screen "41 BWT Ops" 1280x800, template "Template"
   TextField "Text field_60" at 920,365 size 100x30; Text 'GCU'
   GraphicIOField "Graphic I/O field_4" at 920,395 size 100x90; PictureList "GCU"
      ProcessValue <- "100_GCU_AUTO_SEQ_DB_RNG"
   TextField "Text field_70" at 930,485 size 80x25; Text 'Disabled'
   TextField "Text field_71" at 930,485 size 80x25; Text 'Enabled'
      Visibility <- "100_GCU_AUTO_SEQ_DB_RNG"
   Button "Button_4" at 910,355 size 120x170; TextOff 'Text'
      on Release: ActivateScreen("Inert Gas Conditioning Plant", 0)
   TextField "Text field_65" at 730,365 size 100x30; Text 'PGC'
   TextField "Text field_75" at 740,485 size 80x25; Text 'Disabled'
   TextField "Text field_76" at 740,485 size 80x25; Text 'Enabled'
      Visibility <- "10_DI_DATA_E_400_RUN"
   GraphicView "Graphic view_76" at 730,395 size 100x90; Picture "Graphic_251"
   Button "Button_6" at 720,355 size 120x170; TextOff 'Text'
      on Release: ActivateScreen("PGC System", 0)
   TextField "Text field_74" at 1110,365 size 100x30; Text 'IGGS'
   GraphicIOField "Graphic I/O field_1" at 1110,395 size 100x90; PictureList "IGGS"
      ProcessValue <- "14_DQ_Data_24PF1"
   TextField "Text field_62" at 1120,485 size 80x25; Text 'Disabled'
   TextField "Text field_77" at 1120,485 size 80x25; Text 'Enabled'
      Visibility <- "14_DQ_Data_24PF1"
   Button "Button_8" at 1100,355 size 120x170; TextOff 'Text'
      on Release: ActivateScreen("Inert Gas Generator Plant", 0)
   Circle "Circle_1" at 170,240 size 20x20
      Appearance <- "20_TANKS_IP_DATA_RIO_02_FIRST_TANK_BWT_LEVEL_HIHI"
   TextField "Text field_4" at 90,240 size 75x20; Text 'LS422-2P'
   GraphicView "Graphic view_13" at 441,293 size 50x50; Picture "valvevert"
   GraphicView "Graphic view_59" at 199,433 size 518x14; Picture "Graphic_151"
   GraphicView "Logo" at 1,1 size 219x60; Picture "Logo of IGG HMI"
   Button "HmiScreenItemData_1" at 1,50 size 150x43; TextOn 'Back'; TextOff 'Main Index'
      on Release: ActivateScreen("02 Main Index", 0)
   Button "HmiScreenItemData_2" at 1128,64 size 150x43; TextOn 'Back'; TextOff 'BWT Setup'
      on Release: ActivateScreen("Balast Water Treatment Setup", 0)
   DateTimeField "HmiScreenItemData_17" at 1175,0 size 105x30
   DateTimeField "HmiScreenItemData" at 1175,30 size 105x30
   AlarmView "Alarm view_1" at 0,777 size 1280x23
   TextField "Text field_1" at 324,55 size 640x35; Text 'BASIC BARGE TWO TANK CONTROL SYSTEM'
   TextField "Text field_2" at 484,85 size 320x35; Text 'BTCS ENABLED'
      Visibility <- "80_From_HMI_RUN_BTCS"
   TextField "Text field_3" at 484,85 size 320x35; Text 'BTCS DISABLED'
      Visibility <- "80_From_HMI_RUN_BTCS"
   Button "HmiScreenItemData_19" at 700,128 size 570x30; TextOn 'Back'; TextOff 'IGG STEP'; TextList "STEP LIST BTCS"
      ProcessValue <- "2110_BTCS_CNTRL_DB_BTCS_STEP"
   IOField "I/O field_15" at 600,128 size 90x30; Authorization "Commissioning"; FormatPattern 999; Unit  Step
      ProcessValue <- "2110_BTCS_CNTRL_DB_BTCS_STEP"
   Button "HmiScreenItemData_9" at 490,128 size 100x30; TextOn 'Back'; TextOff 'BTCS PLC'
   Button "HmiScreenItemData_3" at 700,168 size 570x30; TextOn 'Back'; TextOff 'IGG STEP'; TextList "STATE LIST BTCS"
      ProcessValue <- "2110_BTCS_CNTRL_DB_BTCS_STATE"
   IOField "I/O field_16" at 600,168 size 90x30; Authorization "Commissioning"; FormatPattern 9; Unit  State
      ProcessValue <- "2110_BTCS_CNTRL_DB_BTCS_STATE"
   Group "Group" at 1100,355 size 120x170; PictureList "IGGS"
   Group "Group_1" at 910,355 size 120x170; PictureList "GCU"
   Group "Group_2" at 720,355 size 120x170; Picture "Graphic_251"
   GraphicView "Graphic view_3" at 506,400 size 50x50; Picture "Graphic_288"
   GraphicView "Graphic view_6" at 346,400 size 50x50; Picture "Graphic_288"
   GraphicView "Graphic view_9" at 615,400 size 50x50; Picture "Graphic_288"
   TextField "Text field_7" at 610,452 size 60x20; Text 'CV-406'
   TextField "Text field_33" at 610,370 size 60x25; Text 'Closed'
      Visibility <- "10_DI_DATA_CV406_CLSD"
   TextField "Text field_14" at 610,370 size 60x25; Text 'Opened'
      Visibility <- "10_DI_DATA_CV406_OPN"
   TextField "Text field_45" at 501,370 size 60x25; Text 'Closed'
      Visibility <- "10_DI_DATA_CV407_CLSD"
   TextField "Text field_11" at 501,370 size 60x25; Text 'Opened'
      Visibility <- "10_DI_DATA_CV407_OPN"
   TextField "Text field_9" at 341,370 size 60x25; Text 'Closed'
      Visibility <- "10_DI_DATA_CV411_CLSD"
   TextField "Text field_10" at 341,370 size 60x25; Text 'Opened'
      Visibility <- "10_DI_DATA_CV411_OPN"
   TextField "Text field_13" at 470,268 size 60x25; Text 'Opened'
      Visibility <- "10_DI_DATA_CV409_OPN"
   TextField "Text field_12" at 470,268 size 60x25; Text 'Closed'
      Visibility <- "10_DI_DATA_CV409_CLSD"
   TextField "Text field_15" at 456,343 size 60x20; Text 'CV-409'
   TextField "Text field_16" at 501,452 size 60x20; Text 'CV-407'
   GraphicView "Graphic view_106" at 444,337 size 14x101; Picture "Graphic_147"
   TextField "Text field_17" at 341,452 size 60x20; Text 'CV-411'
   GraphicView "Graphic view_14" at 444,255 size 14x40; Picture "Graphic_147"
   TextField "Text field_5" at 237,335 size 60x25; Text 'Opened'
      Visibility <- "20_TANKS_IP_DATA_RIO_02_FIRST_TANK_GTT_ISOL_VALVE_OPEN"
   TextField "Text field_6" at 237,335 size 60x25; Text 'Closed'
      Visibility <- "20_TANKS_IP_DATA_RIO_02_FIRST_TANK_GTT_ISOL_VALVE_CLSD"
   TextField "Text field_8" at 238,456 size 60x25; Text 'Opened'
      Visibility <- "20_TANKS_IP_DATA_RIO_02_SECOND_TANK_GTT_ISOL_VALVE_OPEN"
   TextField "Text field_18" at 238,456 size 60x25; Text 'Closed'
      Visibility <- "20_TANKS_IP_DATA_RIO_02_SECOND_TANK_GTT_ISOL_VALVE_CLSD"
   GraphicView "Graphic view_15" at 208,360 size 50x50; Picture "valvevert"
   TextField "Text field_21" at 223,410 size 80x20; Text 'CV-422-2P'
   GraphicView "Graphic view_16" at 211,320 size 14x42; Picture "Graphic_147"
   GraphicView "Graphic view_17" at 209,481 size 50x50; Picture "valvevert"
   TextField "Text field_22" at 224,531 size 80x20; Text 'CV-421-2S'
   GraphicView "Graphic view_18" at 212,405 size 14x79; Picture "Graphic_147"
   GraphicView "Graphic view_11" at 212,527 size 14x33; Picture "Graphic_147"
   Button "Button_1" at 40,130 size 200x150; TextOff 'Tank - 2P'
      Appearance <- "2110_BTCS_CNTRL_DB_PORT_TANK_STS"
   GraphicView "Graphic view_1" at 200,140 size 30x130; Picture "Graphic_183"
   GraphicView "Graphic view_10" at 50,140 size 30x130; Picture "Graphic_183"
   Button "Button_2" at 90,140 size 100x30; TextOff 'Enable / Disable'; TextList "ENBL_DSBL"
      on Press: InvertBit("2110_BTCS_CNTRL_DB_PORT_TANK_STS")
      Appearance <- "2110_BTCS_CNTRL_DB_PORT_TANK_STS"
      ProcessValue <- "2110_BTCS_CNTRL_DB_PORT_TANK_STS"
   Group "Group_3" at 90,240 size 100x20
   Button "Button_7" at 40,600 size 200x150; TextOff 'Tank - 2S'
      Appearance <- "2110_BTCS_CNTRL_DB_STBD_TANK_STS"
   GraphicView "Graphic view_12" at 200,610 size 30x130; Picture "Graphic_183"
   GraphicView "Graphic view_19" at 50,610 size 30x130; Picture "Graphic_183"
   Button "Button_9" at 90,710 size 100x30; TextOff 'Enable / Disable'; TextList "ENBL_DSBL"
      on Press: InvertBit("2110_BTCS_CNTRL_DB_STBD_TANK_STS")
      ProcessValue <- "2110_BTCS_CNTRL_DB_PORT_TANK_STS"
      Appearance <- "2110_BTCS_CNTRL_DB_STBD_TANK_STS"
   Group "Group_4" at 90,615 size 100x20
   TextField "Text field_37" at 5,550 size 90x20; Text 'FIT417 USD'
   IOField "I/O field_10" at 5,570 size 120x25; FormatPattern 9999.9; Unit Nm³/hr
      ProcessValue <- "20_TANKS_IP_DATA_RIO_02_SECOND_TANK_USD_FLOW"
   TextField "Text field_38" at 280,570 size 90x20; Text 'FIT419 MBG'
   IOField "I/O field_11" at 158,570 size 120x25; FormatPattern 9999.9; Unit Nm³/hr
      ProcessValue <- "20_TANKS_IP_DATA_RIO_02_SECOND_TANK_MBG_FLOW"
   TextField "Text field_30" at 5,315 size 90x20; Text 'FIT418 USD'
   IOField "I/O field_5" at 5,290 size 120x25; FormatPattern 9999.9; Unit Nm³/hr
      ProcessValue <- "20_TANKS_IP_DATA_RIO_02_FIRST_TANK_USD_FLOW"
   TextField "Text field_31" at 280,290 size 90x20; Text 'FIT420 MBG'
   IOField "I/O field_6" at 158,290 size 120x25; FormatPattern 9999.9; Unit Nm³/hr
      ProcessValue <- "20_TANKS_IP_DATA_RIO_02_FIRST_TANK_MBG_FLOW"
   IOField "I/O field_30" at 105,355 size 72x25; FormatPattern s999.9; Unit %
      ProcessValue <- "20_TANKS_IP_DATA_RIO_02_FIRST_TANK_BWT_LEVEL"
   IOField "I/O field_31" at 105,483 size 72x25; FormatPattern s999.9; Unit %
      ProcessValue <- "20_TANKS_IP_DATA_RIO_02_SECOND_TANK_BWT_LEVEL"
   IOField "I/O field_32" at 23,355 size 72x25; FormatPattern 999; Unit  DegC
      ProcessValue <- "20_TANKS_IP_DATA_RIO_02_FIRST_TANK_BWT_TEMP"
   IOField "I/O field_33" at 23,483 size 72x25; FormatPattern 999; Unit  DegC
      ProcessValue <- "20_TANKS_IP_DATA_RIO_02_SECOND_TANK_BWT_TEMP"
   IOField "I/O field_34" at 105,386 size 72x25; FormatPattern 9.9; Unit  ph
      ProcessValue <- "20_TANKS_IP_DATA_RIO_02_FIRST_TANK_BWT_PH"
   IOField "I/O field_35" at 105,515 size 72x25; FormatPattern 9.9; Unit  ph
      ProcessValue <- "20_TANKS_IP_DATA_RIO_02_SECOND_TANK_BWT_PH"
   IOField "I/O field_36" at 23,386 size 72x25; FormatPattern 99.9; Unit  mg/l
      ProcessValue <- "20_TANKS_IP_DATA_RIO_02_FIRST_TANK_BWT_DO"
   IOField "I/O field_37" at 23,515 size 72x25; FormatPattern 99.9; Unit  mg/l
      ProcessValue <- "20_TANKS_IP_DATA_RIO_02_SECOND_TANK_BWT_DO"
   IOField "I/O field_2" at 595,481 size 81x25; FormatPattern 999.9; Unit  Barg
      ProcessValue <- "20_TANKS_IP_DATA_RIO_02_FIRST_TANK_DECK_IG_PRESS"
   Button "HmiScreenItemData_4" at 321,635 size 226x75; TextOn 'Back'; TextOff 'MEA Tank Changeover'; TextList "PGC Commissioning"
      on Release: SetBit("PGC_COMMISSION_MODE_DB_Active")
      ProcessValue <- "PGC_COMMISSION_MODE_DB_Button Control"
      Visibility <- "10_DI_DATA_E_400_RUN"
   Circle "Circle_2" at 170,615 size 20x20
      Appearance <- "20_TANKS_IP_DATA_RIO_02_SECOND_TANK_BWT_LEVEL_HIHI"
   TextField "Text field_19" at 90,615 size 75x20; Text 'LS422-2S'

screen "42 BWT Setup" 1280x800, template "Template"
   Button "HmiScreenItemData_1" at 1,1 size 150x43; TextOn 'Back'; TextOff 'Main Index'
      on Release: ActivateScreen("02 Main Index", 0)
   Button "HmiScreenItemData_3" at 1129,1 size 150x43; TextOn 'I&A Compressor Ok'; TextOff 'Back'
      on Release: function_efd93a16()
   AlarmView "Alarm view_1" at 0,777 size 1280x23
   Group "Group_5" at 640,205 size 480x40
   Group "Group_6" at 640,295 size 480x40
   TextField "Text field_31" at 1005,150 size 120x30; Text 'SETUP'
   Button "HmiScreenItemData_19" at 700,60 size 570x30; TextOn 'Back'; TextOff 'IGG STEP'; TextList "STEP LIST BTCS"
      ProcessValue <- "2110_BTCS_CNTRL_DB_BTCS_STEP"
   IOField "I/O field_15" at 600,60 size 90x30; Authorization "Commissioning"; FormatPattern 999; Unit  Step
      ProcessValue <- "2110_BTCS_CNTRL_DB_BTCS_STEP"
   Button "HmiScreenItemData_9" at 490,60 size 100x30; TextOn 'Back'; TextOff 'BTCS PLC'
   Button "HmiScreenItemData_2" at 700,100 size 570x30; TextOn 'Back'; TextOff 'IGG STEP'; TextList "STATE LIST BTCS"
      ProcessValue <- "2110_BTCS_CNTRL_DB_BTCS_STATE"
   IOField "I/O field_16" at 600,100 size 90x30; Authorization "Commissioning"; FormatPattern 9; Unit  State
      ProcessValue <- "2110_BTCS_CNTRL_DB_BTCS_STATE"
   SymbolicIOField "Symbolic I/O field_3" at 360,450 size 140x30; TextOn '1'; TextOff '0'; TextList "Port Tank"
      ProcessValue <- "2110_BTCS_CNTRL_DB_PORT_TANK_STS"
   TextField "Text field_35" at 1025,440 size 100x30; Text 'TANKS'
   SymbolicIOField "Symbolic I/O field_4" at 360,490 size 140x30; TextOn '1'; TextOff '0'; TextList "Port Tank"
      ProcessValue <- "2110_BTCS_CNTRL_DB_STBD_TANK_STS"
   TextField "Text field_37" at 515,450 size 60x30; Text 'O2 :'
   IOField "I/O field_20" at 575,450 size 60x30; FormatPattern 99.99
      ProcessValue <- "20_TANKS_IP_DATA_RIO_02_FIRST_TANK_BWT_DO"
   TextField "Text field_36" at 640,450 size 60x30; Text 'ph :'
   IOField "I/O field_19" at 700,450 size 60x30; FormatPattern 99.99
      ProcessValue <- "20_TANKS_IP_DATA_RIO_02_FIRST_TANK_BWT_PH"
   TextField "Text field_38" at 775,450 size 65x30; Text 'Temp :'
   IOField "I/O field_21" at 840,450 size 60x30; FormatPattern 99.99
      ProcessValue <- "20_TANKS_IP_DATA_RIO_02_FIRST_TANK_BWT_TEMP"
   TextField "Text field_39" at 910,450 size 65x30; Text 'Level :'
   IOField "I/O field_22" at 975,450 size 60x30; FormatPattern 99.9
      ProcessValue <- "20_TANKS_IP_DATA_RIO_02_FIRST_TANK_BWT_LEVEL"
   TextField "Text field_40" at 515,490 size 60x30; Text 'O2 :'
   IOField "I/O field_23" at 575,490 size 60x30; FormatPattern 99.99
      ProcessValue <- "20_TANKS_IP_DATA_RIO_02_SECOND_TANK_BWT_DO"
   TextField "Text field_41" at 640,490 size 60x30; Text 'ph :'
   IOField "I/O field_24" at 700,490 size 60x30; FormatPattern 99.99
      ProcessValue <- "20_TANKS_IP_DATA_RIO_02_SECOND_TANK_BWT_PH"
   TextField "Text field_42" at 775,490 size 65x30; Text 'Temp :'
   IOField "I/O field_25" at 840,490 size 60x30; FormatPattern 99.99
      ProcessValue <- "20_TANKS_IP_DATA_RIO_02_SECOND_TANK_BWT_TEMP"
   TextField "Text field_43" at 910,490 size 65x30; Text 'Level :'
   IOField "I/O field_26" at 975,490 size 60x30; FormatPattern 99.9
      ProcessValue <- "20_TANKS_IP_DATA_RIO_02_SECOND_TANK_BWT_LEVEL"
   Rectangle "Rectangle_5" at 150,340 size 480x40
      Appearance <- "2102_TIME_CALCS_DB_POST_DWELL_TMR_DN"
   TextField "Text field_16" at 155,345 size 200x30; Text 'Post-Dwell Time :'
   IOField "I/O field_9" at 360,345 size 60x30; FormatPattern 999
      ProcessValue <- "2110_BTCS_CNTRL_DB_POST_DWELL_HRS"
   TextField "Text field_17" at 420,345 size 60x30; Text 'Hours'
   IOField "I/O field_10" at 485,345 size 60x30; FormatPattern 99
      ProcessValue <- "2110_BTCS_CNTRL_DB_POST_DWELL_MINS"
   TextField "Text field_18" at 545,345 size 80x30; Text 'Minutes'
   Rectangle "Rectangle_4" at 150,295 size 480x40
      Appearance <- "2102_TIME_CALCS_DB_RE_OX_TMR_DN"
   TextField "Text field_13" at 155,300 size 200x30; Text 'Re-Oxygenate Time :'
   IOField "I/O field_7" at 360,300 size 60x30; FormatPattern 999
      ProcessValue <- "2110_BTCS_CNTRL_DB_RE_OX_HRS"
   TextField "Text field_14" at 420,300 size 60x30; Text 'Hours'
   IOField "I/O field_8" at 485,300 size 60x30; FormatPattern 99
      ProcessValue <- "2110_BTCS_CNTRL_DB_RE_OX_MINS"
   TextField "Text field_15" at 545,300 size 80x30; Text 'Minutes'
   Rectangle "Rectangle_3" at 150,250 size 480x40
      Appearance <- "2102_TIME_CALCS_DB_DWELL_TMR_DN"
   TextField "Text field_10" at 155,255 size 200x30; Text 'Dwell Time :'
   IOField "I/O field_5" at 360,255 size 60x30; FormatPattern 999
      ProcessValue <- "2110_BTCS_CNTRL_DB_DWELL_HRS"
   TextField "Text field_11" at 420,255 size 60x30; Text 'Hours'
   IOField "I/O field_6" at 485,255 size 60x30; FormatPattern 99
      ProcessValue <- "2110_BTCS_CNTRL_DB_DWELL_MINS"
   TextField "Text field_12" at 545,255 size 80x30; Text 'Minutes'
   Rectangle "Rectangle_2" at 150,205 size 480x40
      Appearance <- "2102_TIME_CALCS_DB_DE_OX_TMR_DN"
   TextField "Text field_7" at 155,210 size 200x30; Text 'De-Oxygenate Time :'
   IOField "I/O field_3" at 360,210 size 60x30; FormatPattern 999
      ProcessValue <- "2110_BTCS_CNTRL_DB_DE_OX_HRS"
   TextField "Text field_8" at 420,210 size 60x30; Text 'Hours'
   IOField "I/O field_4" at 485,210 size 60x30; FormatPattern 99
      ProcessValue <- "2110_BTCS_CNTRL_DB_DE_OX_MINS"
   TextField "Text field_9" at 545,210 size 80x30; Text 'Minutes'
   Rectangle "Rectangle_1" at 150,160 size 480x40
      Appearance <- "2102_TIME_CALCS_DB_PRE_DWELL_TMR_DN"
   TextField "Text field_4" at 155,165 size 200x30; Text 'Pre-Dwell Time :'
   IOField "I/O field_1" at 360,165 size 60x30; FormatPattern 999
      ProcessValue <- "2110_BTCS_CNTRL_DB_PRE_DWELL_HRS"
   TextField "Text field_5" at 420,165 size 60x30; Text 'Hours'
   IOField "I/O field_2" at 485,165 size 60x30; FormatPattern 99
      ProcessValue <- "2110_BTCS_CNTRL_DB_PRE_DWELL_MINS"
   TextField "Text field_6" at 545,165 size 80x30; Text 'Minutes'
   Rectangle "Rectangle_6" at 640,205 size 480x40
      Appearance <- "2102_TIME_CALCS_DB_DE_OX_SP_TMR_DN"
   TextField "Text field_19" at 645,210 size 200x30; Text 'At De-Ox Setpoint :'
   IOField "I/O field_11" at 850,210 size 60x30; FormatPattern 999
      ProcessValue <- "2110_BTCS_CNTRL_DB_DE_OX_SP_HRS"
   TextField "Text field_20" at 910,210 size 60x30; Text 'Hours'
   IOField "I/O field_12" at 975,210 size 60x30; FormatPattern 99
      ProcessValue <- "2110_BTCS_CNTRL_DB_DE_OX_SP_MINS"
   TextField "Text field_21" at 1035,210 size 80x30; Text 'Minutes'
   Rectangle "Rectangle_7" at 640,295 size 480x40
      Appearance <- "2102_TIME_CALCS_DB_RE_OX_SP_TMR_DN"
   TextField "Text field_22" at 645,300 size 200x30; Text 'At Re-Ox Setpoint :'
   IOField "I/O field_13" at 850,300 size 60x30; FormatPattern 999
      ProcessValue <- "2110_BTCS_CNTRL_DB_RE_OX_SP_HRS"
   TextField "Text field_23" at 910,300 size 60x30; Text 'Hours'
   IOField "I/O field_14" at 975,300 size 60x30; FormatPattern 99
      ProcessValue <- "2110_BTCS_CNTRL_DB_RE_OX_SP_MINS"
   TextField "Text field_24" at 1035,300 size 80x30; Text 'Minutes'

screen "09 Sys Config" 1280x800, template "Template"
   Circle "Circle_2" at 221,236 size 29x29
      Appearance <- "82_To_HMI_CRNT_MODE_IGG"
   Button "HmiScreenItemData_1" at 1,1 size 150x43; TextOn 'Back'; TextOff 'Main Index'
      on Release: ActivateScreen("02 Main Index", 0)
   Button "HmiScreenItemData_8" at 44,70 size 230x29; TextOn 'Back'; TextOff 'IGG Mode of Operation'
   Circle "Circle_1" at 221,177 size 29x29
      Appearance <- "82_To_HMI_CRNT_MODE_IGG"
   Button "HmiScreenItemData_4" at 50,167 size 150x51; TextOn 'Back'; TextOff 'Manual'; Authorization "Operating Mode"
      on Press: function_b14e0dd5("80_From_HMI_Request_Manual(1)", 0)
   Circle "Circle_9" at 221,116 size 29x29
      Appearance <- "82_To_HMI_CRNT_MODE_IGG"
   TextField "Text field_13" at 293,112 size 93x21; Text 'Description'
   IOField "I/O field_13" at 463,189 size 226x30; FormatPattern 9999999999999999999999999999999999999999
      ProcessValue <- "db_time_sync_time_system_READ"
   Button "HmiScreenItemData_26" at 284,70 size 421x29; TextOn 'Back'; TextOff 'Time Setting'
   Button "HmiScreenItemData_24" at 291,231 size 166x30; TextOn 'Back'; TextOff 'Set System Time'; Authorization "Parameter Change"
      on Activate: function_cbf290fd(0, 0)
   Button "HmiScreenItemData_16" at 894,69 size 187x29; TextOn 'Back'; TextOff 'IO'
   Button "HmiScreenItemData_2" at 719,69 size 163x29; TextOn 'Back'; TextOff 'Runtime'
   Button "HmiScreenItemData_10" at 725,107 size 150x51; TextOn 'Back'; TextOff 'Reset AUTO'; Authorization "User administration"
      on Press: function_b14e0dd5("80_From_HMI_RST_AUT_SEQ(1)", 0)
      Appearance <- "80_From_HMI_RST_AUT_SEQ(1)"
   DateTimeField "Date/time field_1" at 463,231 size 226x30; Authorization "Parameter Change"
   TextField "Text field_14" at 314,195 size 142x20; Text 'System Time (UTC)'
   Button "HmiScreenItemData_23" at 50,106 size 150x51; TextOn 'Back'; TextOff 'Full Automation'; Authorization "Operating Mode"
      on Press: function_b14e0dd5("80_From_HMI_Request_Auto(1)", 0)
   Button "HmiScreenItemData_3" at 1129,1 size 150x43; TextOn 'I&A Compressor Ok'; TextOff 'Back'
      on Release: function_efd93a16()
   Button "HmiScreenItemData_7" at 50,228 size 150x51; TextOn 'Back'; TextOff 'FAT Mode'; Authorization "User administration"
      on Press: InvertBit("80_From_HMI_FAT_Mode"); function_b14e0dd5("80_From_HMI_Request_Auto(1)", 0)
   Button "HmiScreenItemData_11" at 725,232 size 150x51; TextOn 'Back'; TextOff 'IGG Standalone'; Authorization "Operating Mode"
      on Press: InvertBit("80_From_HMI_IGG_STND_ALN")
      Appearance <- "80_From_HMI_IGG_STND_ALN"
   Button "HmiScreenItemData_12" at 910,100 size 150x51; TextOn 'Back'; TextOff 'P301 Present'; TextList "P301 Present"; Authorization "Operating Mode"
      on Press: InvertBit("80_From_HMI_P301_PRSNT(1)")
      Appearance <- "80_From_HMI_P301_PRSNT(1)"
      ProcessValue <- "80_From_HMI_P301_PRSNT(1)"
   Button "HmiScreenItemData_13" at 910,155 size 150x51; TextOn 'Back'; TextOff 'CV312 Present'; TextList "CV312 Present"; Authorization "User administration"
      on Press: InvertBit("80_From_HMI_CV312_PRSNT")
      Appearance <- "80_From_HMI_CV312_PRSNT"
      ProcessValue <- "80_From_HMI_CV312_PRSNT"
   Button "HmiScreenItemData_14" at 910,212 size 150x51; TextOn 'Back'; TextOff 'CV431 Present'; TextList "CV431 Present"; Authorization "Operating Mode"
      on Press: InvertBit("80_From_HMI_CV431_PRSNT")
      Appearance <- "80_From_HMI_CV431_PRSNT"
      ProcessValue <- "80_From_HMI_CV431_PRSNT"
   Button "HmiScreenItemData_15" at 910,269 size 150x51; TextOn 'Back'; TextOff 'CV432 Present'; TextList "CV432 Present"; Authorization "Operating Mode"
      on Press: InvertBit("80_From_HMI_CV432_PRSNT")
      Appearance <- "80_From_HMI_CV432_PRSNT"
      ProcessValue <- "80_From_HMI_CV432_PRSNT"
   Button "HmiScreenItemData_18" at 725,166 size 150x51; TextOn 'Back'; TextOff 'Silence Buzzer'; Authorization "User administration"
      on Press: function_b14e0dd5("80_From_HMI_SLNCE_BZR", 0)
      Appearance <- "80_From_HMI_SLNCE_BZR"
   AlarmView "Alarm view_1" at 0,777 size 1280x23
   IOField "I/O field_9" at 1024,352 size 60x30; Authorization "Commissioning"; FormatPattern 99; Unit  s
      ProcessValue <- "80_From_HMI_Beacon frequency"
   IOField "I/O field_10" at 1025,389 size 60x30; Authorization "Commissioning"; FormatPattern 99; Unit  min
      ProcessValue <- "80_From_HMI_Buzzer reset time"
   TextField "Text field_9" at 895,358 size 138x20; Text 'Beacon frequency'
   TextField "Text field_10" at 895,394 size 100x20; Text 'Buzzer reset'

screen "07 BWTS MAIN" 1280x800, template "Template"
   Rectangle "Rectangle_2" at 150,205 size 480x40
      Appearance <- "2102_TIME_CALCS_DB_DE_OX_TMR_DN"
   TextField "Text field_7" at 155,210 size 200x30; Text 'De-Oxygenate Time :'
   IOField "I/O field_3" at 360,210 size 60x30; FormatPattern 999
      ProcessValue <- "2110_BTCS_CNTRL_DB_DE_OX_HRS"
   TextField "Text field_8" at 420,210 size 60x30; Text 'Hours'
   IOField "I/O field_4" at 485,210 size 60x30; FormatPattern 99
      ProcessValue <- "2110_BTCS_CNTRL_DB_DE_OX_MINS"
   TextField "Text field_9" at 545,210 size 80x30; Text 'Minutes'
   Rectangle "Rectangle_3" at 150,250 size 480x40
      Appearance <- "2102_TIME_CALCS_DB_DWELL_TMR_DN"
   TextField "Text field_10" at 155,255 size 200x30; Text 'Dwell Time :'
   IOField "I/O field_5" at 360,255 size 60x30; FormatPattern 999
      ProcessValue <- "2110_BTCS_CNTRL_DB_DWELL_HRS"
   TextField "Text field_11" at 420,255 size 60x30; Text 'Hours'
   IOField "I/O field_6" at 485,255 size 60x30; FormatPattern 99
      ProcessValue <- "2110_BTCS_CNTRL_DB_DWELL_MINS"
   TextField "Text field_12" at 545,255 size 80x30; Text 'Minutes'
   Rectangle "Rectangle_4" at 150,295 size 480x40
      Appearance <- "2102_TIME_CALCS_DB_RE_OX_TMR_DN"
   TextField "Text field_13" at 155,300 size 200x30; Text 'Re-Oxygenate Time :'
   IOField "I/O field_7" at 360,300 size 60x30; FormatPattern 999
      ProcessValue <- "2110_BTCS_CNTRL_DB_RE_OX_HRS"
   TextField "Text field_14" at 420,300 size 60x30; Text 'Hours'
   IOField "I/O field_8" at 485,300 size 60x30; FormatPattern 99
      ProcessValue <- "2110_BTCS_CNTRL_DB_RE_OX_MINS"
   TextField "Text field_15" at 545,300 size 80x30; Text 'Minutes'
   Rectangle "Rectangle_5" at 150,340 size 480x40
      Appearance <- "2102_TIME_CALCS_DB_POST_DWELL_TMR_DN"
   TextField "Text field_16" at 155,345 size 200x30; Text 'Post-Dwell Time :'
   IOField "I/O field_9" at 360,345 size 60x30; FormatPattern 999
      ProcessValue <- "2110_BTCS_CNTRL_DB_POST_DWELL_HRS"
   TextField "Text field_17" at 420,345 size 60x30; Text 'Hours'
   IOField "I/O field_10" at 485,345 size 60x30; FormatPattern 99
      ProcessValue <- "2110_BTCS_CNTRL_DB_POST_DWELL_MINS"
   TextField "Text field_18" at 545,345 size 80x30; Text 'Minutes'
   Rectangle "Rectangle_6" at 640,205 size 480x40
      Appearance <- "2102_TIME_CALCS_DB_DE_OX_SP_TMR_DN"
   TextField "Text field_19" at 645,210 size 200x30; Text 'At De-Ox Setpoint :'
   IOField "I/O field_11" at 850,210 size 60x30; FormatPattern 999
      ProcessValue <- "2110_BTCS_CNTRL_DB_DE_OX_SP_HRS"
   TextField "Text field_20" at 910,210 size 60x30; Text 'Hours'
   IOField "I/O field_12" at 975,210 size 60x30; FormatPattern 99
      ProcessValue <- "2110_BTCS_CNTRL_DB_DE_OX_SP_MINS"
   TextField "Text field_21" at 1035,210 size 80x30; Text 'Minutes'
   Rectangle "Rectangle_7" at 640,295 size 480x40
      Appearance <- "2102_TIME_CALCS_DB_RE_OX_SP_TMR_DN"
   TextField "Text field_22" at 645,300 size 200x30; Text 'At Re-Ox Setpoint :'
   IOField "I/O field_13" at 850,300 size 60x30; FormatPattern 999
      ProcessValue <- "2110_BTCS_CNTRL_DB_RE_OX_SP_HRS"
   TextField "Text field_23" at 910,300 size 60x30; Text 'Hours'
   IOField "I/O field_14" at 975,300 size 60x30; FormatPattern 99
      ProcessValue <- "2110_BTCS_CNTRL_DB_RE_OX_SP_MINS"
   TextField "Text field_24" at 1035,300 size 80x30; Text 'Minutes'
   TextField "Text field_25" at 155,435 size 200x30; Text 'Total Sequence Time:'
   IOField "I/O field_15" at 360,435 size 60x30; FormatPattern 999
      ProcessValue <- "2110_BTCS_CNTRL_DB_TOT_SEQ_HRS"
   TextField "Text field_26" at 420,435 size 60x30; Text 'Hours'
   IOField "I/O field_16" at 485,435 size 60x30; FormatPattern 99
      ProcessValue <- "2110_BTCS_CNTRL_DB_TOT_SEQ_MINS"
   TextField "Text field_27" at 545,435 size 80x30; Text 'Minutes'
   TextField "Text field_28" at 155,625 size 200x30; Text 'Remaining Time:'
   IOField "I/O field_17" at 360,625 size 60x30; FormatPattern 999
      ProcessValue <- "2110_BTCS_CNTRL_DB_RMNG_SEQ_HRS"
   TextField "Text field_29" at 420,625 size 60x30; Text 'Hours'
   IOField "I/O field_18" at 485,625 size 60x30; FormatPattern 99
      ProcessValue <- "2110_BTCS_CNTRL_DB_RMNG_SEQ_MINS"
   TextField "Text field_30" at 545,625 size 80x30; Text 'Minutes'
   Button "HmiScreenItemData_1" at 10,10 size 160x50; TextOn 'Back'; TextOff 'Main Index'
      on Release: ActivateScreen("02 Main Index", 0)
   TextField "Text field_1" at 320,10 size 640x35; Text 'BASIC BARGE TWO TANK CONTROL SYSTEM'
   Button "HmiScreenItemData_2" at 1110,10 size 160x50; TextOn 'Back'; TextOff 'Enable'
      on Press: ResetBit("80_From_HMI_RUN_BWTS"); SetBit("80_From_HMI_RUN_BTCS")
      Visibility <- "80_From_HMI_RUN_BWTS"
   Button "HmiScreenItemData_3" at 918,75 size 160x50; TextOn 'Back'; TextOff 'Disable'
      on Press: ResetBit("80_From_HMI_RUN_BTCS"); SetBit("80_From_HMI_RUN_BWTS")
      Visibility <- "80_From_HMI_RUN_BTCS"
   TextField "Text field_2" at 480,40 size 320x35; Text 'BTCS ENABLED'
      Visibility <- "80_From_HMI_RUN_BTCS"
   TextField "Text field_3" at 480,40 size 320x35; Text 'BTCS DISABLED'
      Visibility <- "80_From_HMI_RUN_BTCS"
   Button "Button_2" at 10,70 size 160x50; TextOn 'User Account'; TextOff 'Alarm Log'; Authorization "User administration"
      on Release: ActivateScreen("04 Alarm Log", 0)
   Group "Group_1" at 150,205 size 480x40
   Group "Group_2" at 150,250 size 480x40
   Group "Group_3" at 150,295 size 480x40
   Group "Group_4" at 150,340 size 480x40
   Group "Group_5" at 640,205 size 480x40
   Group "Group_6" at 640,295 size 480x40
   Group "Group_7" at 150,430 size 480x40
   Group "Group_8" at 150,620 size 480x40
   TextField "Text field_31" at 1005,150 size 120x30; Text 'SETUP'
   TextField "Text field_32" at 1005,420 size 120x30; Text 'CONTROL'
   Button "Button_1" at 150,520 size 230x50; TextOff 'ACCEPT & LAUNCH'
      on Release: ResetBit("2110_BTCS_CNTRL_DB_START_SEQ")
      on Press: SetBit("2110_BTCS_CNTRL_DB_START_SEQ")
      Appearance <- "2110_BTCS_CNTRL_DB_BTCS_STATE"
      Visibility <- "2102_TIME_CALCS_DB_TIMES_VALID"
   SymbolicIOField "Symbolic I/O field_1" at 640,480 size 480x30; TextOn '1'; TextOff '0'; TextList "STATE LIST BTCS"
      ProcessValue <- "2110_BTCS_CNTRL_DB_BTCS_STATE"
   TextField "Text field_33" at 150,480 size 480x35; Text 'TIMES NOT VALID'
      Visibility <- "2102_TIME_CALCS_DB_TIMES_VALID"
   TextField "Text field_34" at 150,480 size 480x35; Text 'TIMES VALID'
      Visibility <- "2102_TIME_CALCS_DB_TIMES_VALID"
   SymbolicIOField "Symbolic I/O field_2" at 640,580 size 480x30; TextOn '1'; TextOff '0'; TextList "STEP LIST BTCS"
      ProcessValue <- "2110_BTCS_CNTRL_DB_BTCS_STEP"
   Button "HmiScreenItemData_4" at 1110,70 size 160x50; TextOn 'Back'; TextOff 'Master Reset'
      on Press: ResetBit("2110_BTCS_CNTRL_DB_RESET_ALL"); SetBit("2110_BTCS_CNTRL_DB_RESET_ALL")
      Visibility <- "80_From_HMI_RUN_BTCS"
   SymbolicIOField "Symbolic I/O field_3" at 360,700 size 140x30; TextOn '1'; TextOff '0'; TextList "Port Tank"
      ProcessValue <- "2110_BTCS_CNTRL_DB_PORT_TANK_STS"
   Button "Button_4" at 150,700 size 180x30; TextOff 'Port Tank'
      on Press: InvertBit("2110_BTCS_CNTRL_DB_PORT_TANK_STS")
      Appearance <- "2110_BTCS_CNTRL_DB_PORT_TANK_STS"
   TextField "Text field_35" at 1025,690 size 100x30; Text 'TANKS'
   SymbolicIOField "Symbolic I/O field_4" at 360,740 size 140x30; TextOn '1'; TextOff '0'; TextList "Port Tank"
      ProcessValue <- "2110_BTCS_CNTRL_DB_STBD_TANK_STS"
   Button "Button_5" at 150,740 size 180x30; TextOff 'Starboard Tank'
      on Press: InvertBit("2110_BTCS_CNTRL_DB_STBD_TANK_STS")
      Appearance <- "2110_BTCS_CNTRL_DB_STBD_TANK_STS"
   TextField "Text field_37" at 515,700 size 60x30; Text 'O2 :'
   IOField "I/O field_20" at 575,700 size 60x30; FormatPattern 99.99
      ProcessValue <- "20_TANKS_IP_DATA_RIO_02_FIRST_TANK_BWT_DO"
   TextField "Text field_36" at 640,700 size 60x30; Text 'ph :'
   IOField "I/O field_19" at 700,700 size 60x30; FormatPattern 99.99
      ProcessValue <- "20_TANKS_IP_DATA_RIO_02_FIRST_TANK_BWT_PH"
   TextField "Text field_38" at 775,700 size 65x30; Text 'Temp :'
   IOField "I/O field_21" at 840,700 size 60x30; FormatPattern 99.99
      ProcessValue <- "20_TANKS_IP_DATA_RIO_02_FIRST_TANK_BWT_TEMP"
   TextField "Text field_39" at 910,700 size 65x30; Text 'Level :'
   IOField "I/O field_22" at 975,700 size 60x30; FormatPattern 99.9
      ProcessValue <- "20_TANKS_IP_DATA_RIO_02_FIRST_TANK_BWT_LEVEL"
   TextField "Text field_40" at 515,740 size 60x30; Text 'O2 :'
   IOField "I/O field_23" at 575,740 size 60x30; FormatPattern 99.99
      ProcessValue <- "20_TANKS_IP_DATA_RIO_02_SECOND_TANK_BWT_DO"
   TextField "Text field_41" at 640,740 size 60x30; Text 'ph :'
   IOField "I/O field_24" at 700,740 size 60x30; FormatPattern 99.99
      ProcessValue <- "20_TANKS_IP_DATA_RIO_02_SECOND_TANK_BWT_PH"
   TextField "Text field_42" at 775,740 size 65x30; Text 'Temp :'
   IOField "I/O field_25" at 840,740 size 60x30; FormatPattern 99.99
      ProcessValue <- "20_TANKS_IP_DATA_RIO_02_SECOND_TANK_BWT_TEMP"
   TextField "Text field_43" at 910,740 size 65x30; Text 'Level :'
   IOField "I/O field_26" at 975,740 size 60x30; FormatPattern 99.9
      ProcessValue <- "20_TANKS_IP_DATA_RIO_02_SECOND_TANK_BWT_LEVEL"
   Group "Group" at 150,160 size 480x40
   Group "Group_9" at 150,160 size 480x40
   Group "Group_10" at 150,340 size 480x40
   Group "Group_12" at 150,295 size 480x40
   Group "Group_13" at 640,205 size 480x40
   Group "Group_14" at 150,250 size 480x40
   Group "Group_15" at 150,205 size 480x40
   Group "Group_16" at 640,295 size 480x40
   Rectangle "Rectangle_15" at 150,480 size 480x130
      Visibility <- "2100_AUTO_SEQ_DB_SEQ_RNG"
   Button "Button_3" at 400,520 size 230x50; TextOff 'ABORT - STOP'
      on Release: ResetBit("2110_BTCS_CNTRL_DB_STOP_SEQ")
      on Press: SetBit("2110_BTCS_CNTRL_DB_STOP_SEQ")
      Appearance <- "2110_BTCS_CNTRL_DB_BTCS_STATE"
   TextField "Text field_48" at 23,309 size 1188x123; Text 'Re - Work Required Througout This page'
   Rectangle "Rectangle_1" at 150,160 size 480x40
      Appearance <- "2102_TIME_CALCS_DB_PRE_DWELL_TMR_DN"
   TextField "Text field_4" at 155,165 size 200x30; Text 'Pre-Dwell Time :'
   IOField "I/O field_1" at 360,165 size 60x30; FormatPattern 999
      ProcessValue <- "2110_BTCS_CNTRL_DB_PRE_DWELL_HRS"
   TextField "Text field_5" at 420,165 size 60x30; Text 'Hours'
   IOField "I/O field_2" at 485,165 size 60x30; FormatPattern 99
      ProcessValue <- "2110_BTCS_CNTRL_DB_PRE_DWELL_MINS"
   TextField "Text field_6" at 545,165 size 80x30; Text 'Minutes'
   Rectangle "Rectangle_13" at 150,160 size 480x40
      Visibility <- "2100_AUTO_SEQ_DB_SEQ_RNG"
      Appearance <- "2102_TIME_CALCS_DB_PRE_DWELL_TMR_DN"
   TextField "Text field_44" at 155,165 size 310x30; Text 'Pre-Dwell Time Remaining :'
      Visibility <- "2100_AUTO_SEQ_DB_SEQ_RNG"
   IOField "I/O field_28" at 465,165 size 80x30; FormatPattern 999999
      Visibility <- "2100_AUTO_SEQ_DB_SEQ_RNG"
      ProcessValue <- "2102_TIME_CALCS_DB_PRE_DWELL_MINS_RMNG"
   TextField "Text field_46" at 545,165 size 80x30; Text 'Minutes'
      Visibility <- "2100_AUTO_SEQ_DB_SEQ_RNG"
   Rectangle "Rectangle_14" at 150,340 size 480x40
      Visibility <- "2100_AUTO_SEQ_DB_SEQ_RNG"
      Appearance <- "2102_TIME_CALCS_DB_POST_DWELL_TMR_DN"
   TextField "Text field_45" at 155,345 size 310x30; Text 'Post-Dwell Time Remaining :'
      Visibility <- "2100_AUTO_SEQ_DB_SEQ_RNG"
   IOField "I/O field_27" at 465,345 size 80x30; FormatPattern 999999
      ProcessValue <- "2102_TIME_CALCS_DB_POST_DWELL_MINS_RMNG"
      Visibility <- "2100_AUTO_SEQ_DB_SEQ_RNG"
   TextField "Text field_47" at 545,345 size 80x30; Text 'Minutes'
      Visibility <- "2100_AUTO_SEQ_DB_SEQ_RNG"
   Rectangle "Rectangle_16" at 150,295 size 480x40
      Visibility <- "2100_AUTO_SEQ_DB_SEQ_RNG"
      Appearance <- "2102_TIME_CALCS_DB_RE_OX_TMR_DN"
   TextField "Text field_50" at 155,300 size 310x30; Text 'Re-Oxygenate Time Remaining :'
      Visibility <- "2100_AUTO_SEQ_DB_SEQ_RNG"
   IOField "I/O field_30" at 465,300 size 80x30; FormatPattern 999999
      ProcessValue <- "2102_TIME_CALCS_DB_RE_OX_MINS_RMNG"
      Visibility <- "2100_AUTO_SEQ_DB_SEQ_RNG"
   TextField "Text field_51" at 545,300 size 80x30; Text 'Minutes'
      Visibility <- "2100_AUTO_SEQ_DB_SEQ_RNG"
   Rectangle "Rectangle_17" at 640,205 size 480x40
      Visibility <- "2100_AUTO_SEQ_DB_SEQ_RNG"
      Appearance <- "2102_TIME_CALCS_DB_DE_OX_SP_TMR_DN"
   TextField "Text field_52" at 645,210 size 310x30; Text 'At De-Ox Time Remaining :'
      Visibility <- "2100_AUTO_SEQ_DB_SEQ_RNG"
   IOField "I/O field_31" at 955,210 size 80x30; FormatPattern 999999
      ProcessValue <- "2102_TIME_CALCS_DB_DE_OX_SP_MINS_RMNG"
      Visibility <- "2100_AUTO_SEQ_DB_SEQ_RNG"
   TextField "Text field_53" at 1035,210 size 80x30; Text 'Minutes'
      Visibility <- "2100_AUTO_SEQ_DB_SEQ_RNG"
   Rectangle "Rectangle_18" at 150,250 size 480x40
      Visibility <- "2100_AUTO_SEQ_DB_SEQ_RNG"
      Appearance <- "2102_TIME_CALCS_DB_DWELL_TMR_DN"
   TextField "Text field_54" at 155,255 size 310x30; Text 'Dwell Time Remaining :'
      Visibility <- "2100_AUTO_SEQ_DB_SEQ_RNG"
   IOField "I/O field_32" at 465,255 size 80x30; FormatPattern 999999
      ProcessValue <- "2102_TIME_CALCS_DB_DWELL_MINS_RMNG"
      Visibility <- "2100_AUTO_SEQ_DB_SEQ_RNG"
   TextField "Text field_55" at 545,255 size 80x30; Text 'Minutes'
      Visibility <- "2100_AUTO_SEQ_DB_SEQ_RNG"
   Rectangle "Rectangle_19" at 150,205 size 480x40
      Visibility <- "2100_AUTO_SEQ_DB_SEQ_RNG"
      Appearance <- "2102_TIME_CALCS_DB_DE_OX_TMR_DN"
   TextField "Text field_56" at 155,210 size 310x30; Text 'De-Oxygenate Time Remaining :'
      Visibility <- "2100_AUTO_SEQ_DB_SEQ_RNG"
   IOField "I/O field_33" at 465,210 size 80x30; FormatPattern 999999
      ProcessValue <- "2102_TIME_CALCS_DB_DE_OX_MINS_RMNG"
      Visibility <- "2100_AUTO_SEQ_DB_SEQ_RNG"
   TextField "Text field_57" at 545,210 size 80x30; Text 'Minutes'
      Visibility <- "2100_AUTO_SEQ_DB_SEQ_RNG"
   Rectangle "Rectangle_20" at 640,295 size 480x40
      Visibility <- "2100_AUTO_SEQ_DB_SEQ_RNG"
      Appearance <- "2102_TIME_CALCS_DB_RE_OX_SP_TMR_DN"
   TextField "Text field_58" at 645,300 size 310x30; Text 'At Re-Ox Time Remaining :'
      Visibility <- "2100_AUTO_SEQ_DB_SEQ_RNG"
   IOField "I/O field_34" at 955,300 size 80x30; FormatPattern 999999
      ProcessValue <- "2102_TIME_CALCS_DB_RE_OX_SP_MINS_RMNG"
      Visibility <- "2100_AUTO_SEQ_DB_SEQ_RNG"
   TextField "Text field_59" at 1035,300 size 80x30; Text 'Minutes'
      Visibility <- "2100_AUTO_SEQ_DB_SEQ_RNG"

screen "Inert Gas Conditioning Plant" 1280x800, template "Template_lite"
   on GenerateScreen: "TitleUpdater"()
   GraphicView "Graphic view_20" at 359,634 size 43x62; Picture "Graphic_72"
   GraphicView "Graphic view_52" at 746,80 size 58x108; Picture "Graphic_72"
   GraphicView "Graphic view_63" at 991,218 size 58x108; Picture "Graphic_72"
   GraphicView "Graphic view_64" at 1096,218 size 58x108; Picture "Graphic_72"
   Button "Button_2" at 573,588 size 60x25; TextOn 'Alarm'; TextOff 'OK'
      Appearance <- "10_DI_DATA_P_303_OK"
   TextField "Text field_49" at 573,588 size 60x25; Text 'Enabled'
      Appearance <- "14_DQ_DATA_P_303"
      Visibility <- "14_DQ_DATA_P_303"
   Button "Button_3" at 187,631 size 60x25; TextOn 'Alarm'; TextOff 'OK'
      Appearance <- "10_DI_DATA_P_304_OK"
   TextField "Text field_19" at 187,631 size 60x25; Text 'Enabled'
      Appearance <- "14_DQ_DATA_P_304"
      Visibility <- "14_DQ_DATA_P_304"
   Button "HmiScreenItemData_8" at 228,5 size 355x40; TextOn 'Back'; TextOff 'Text'
   TextField "Screen title" at 214,1 size 373x50; Text 'Screen title'
   Circle "Circle_73" at 594,11 size 10x10
      VerticalMovement <- "E-400 Animation_DB_Animation"
      Visibility <- "10_DI_DATA_E_400_RUN"
   Circle "Circle_45" at 592,89 size 10x10
      VerticalMovement <- "E-400 Animation_DB_Animation"
      Visibility <- "10_DI_DATA_E_400_RUN"
   Circle "Circle_84" at 591,169 size 10x10
      HorizontalMovement <- "E-400 Animation_DB_Animation"
      Visibility <- "10_DI_DATA_E_400_RUN"
   Circle "Circle_26" at 706,169 size 10x10
      Visibility <- "10_DI_DATA_CV406_CLSD"
      HorizontalMovement <- "E-400 Animation_DB_Animation"
   Circle "Circle_27" at 748,169 size 10x10
      Visibility <- "10_DI_DATA_CV406_CLSD"
      HorizontalMovement <- "E-400 Animation_DB_Animation"
   Circle "Circle_28" at 811,169 size 10x10
      Visibility <- "10_DI_DATA_CV407_CLSD"
      HorizontalMovement <- "E-400 Animation_DB_Animation"
   Circle "Circle_29" at 876,169 size 10x10
      Visibility <- "10_DI_DATA_CV407_CLSD"
      HorizontalMovement <- "E-400 Animation_DB_Animation"
   Circle "Circle_72" at 882,168 size 10x10
      Visibility <- "10_DI_DATA_CV407_CLSD"
      HorizontalMovement <- "E-400 Animation_DB_Animation"
   Circle "Circle_30" at 929,168 size 10x10
      Visibility <- "10_DI_DATA_CV407_CLSD"
      HorizontalMovement <- "E-400 Animation_DB_Animation"
   Circle "Circle_71" at 940,168 size 10x10
      Visibility <- "10_DI_DATA_CV407_CLSD"
      HorizontalMovement <- "E-400 Animation_DB_Animation"
   Circle "Circle_31" at 944,304 size 10x10
      Visibility <- "10_DI_DATA_CV407_CLSD"
      VerticalMovement <- "E-400 Animation_DB_Animation"
   Circle "Circle_42" at 995,305 size 10x10
      Visibility <- "10_DI_DATA_CV407_CLSD"
      HorizontalMovement <- "E-400 Animation_DB_Animation"
   Circle "Circle_44" at 1066,143 size 10x10
      Visibility <- "10_DI_DATA_CV409_CLSD"
      VerticalMovement <- "E-400 Animation_DB_Animation"
   Circle "Circle_43" at 1066,224 size 10x10
      Visibility <- "10_DI_DATA_CV409_CLSD"
      VerticalMovement <- "E-400 Animation_DB_Animation"
   Circle "Circle_32" at 1098,306 size 10x10
      Visibility <- "10_DI_DATA_CV411_CLSD"
      HorizontalMovement <- "E-400 Animation_DB_Animation"
   Circle "Circle_82" at 1185,305 size 10x10
      Visibility <- "10_DI_DATA_CV411_CLSD"
      HorizontalMovement <- "E-400 Animation_DB_Animation"
   Circle "Circle_38" at 389,247 size 9x9
      DiagonalMovement <- "E-400 Animation_DB_Animation"
      Visibility <- "10_DI_DATA_E_400_RUN"
   Circle "Circle_57" at 402,247 size 10x10
      DiagonalMovement <- "E-400 Animation_DB_Animation"
      Visibility <- "10_DI_DATA_E_400_RUN"
   Circle "Circle_40" at 417,247 size 10x10
      DiagonalMovement <- "E-400 Animation_DB_Animation"
      Visibility <- "10_DI_DATA_E_400_RUN"
   Circle "Circle_58" at 433,247 size 10x10
      DiagonalMovement <- "E-400 Animation_DB_Animation"
      Visibility <- "10_DI_DATA_E_400_RUN"
   Circle "Circle_60" at 475,162 size 10x10
      DiagonalMovement <- "E-400 Animation_DB_Animation"
      Visibility <- "10_DI_DATA_E_400_RUN"
   Circle "Circle_41" at 474,180 size 10x10
      DiagonalMovement <- "E-400 Animation_DB_Animation"
      Visibility <- "10_DI_DATA_E_400_RUN"
   Circle "Circle_39" at 475,172 size 9x9
      DiagonalMovement <- "E-400 Animation_DB_Animation"
      Visibility <- "10_DI_DATA_E_400_RUN"
   Circle "Circle_59" at 475,152 size 10x10
      DiagonalMovement <- "E-400 Animation_DB_Animation"
      Visibility <- "10_DI_DATA_E_400_RUN"
   Circle "Circle_87" at 448,247 size 10x10
      DiagonalMovement <- "E-400 Animation_DB_Animation"
      Visibility <- "10_DI_DATA_E_400_RUN"
   Circle "Circle_88" at 462,247 size 10x10
      DiagonalMovement <- "E-400 Animation_DB_Animation"
      Visibility <- "10_DI_DATA_E_400_RUN"
   Circle "Circle_89" at 474,190 size 10x10
      DiagonalMovement <- "E-400 Animation_DB_Animation"
      Visibility <- "10_DI_DATA_E_400_RUN"
   Circle "Circle_90" at 474,199 size 10x10
      DiagonalMovement <- "E-400 Animation_DB_Animation"
      Visibility <- "10_DI_DATA_E_400_RUN"
   Circle "Circle_33" at 239,444 size 10x10
      DiagonalMovement <- "E-400 Animation_DB_Animation"
      Visibility <- "10_DI_DATA_E_400_RUN"
   Circle "Circle_34" at 240,306 size 11x11
      Visibility <- "10_DI_DATA_E_400_RUN"
      VerticalMovement <- "E-400 Animation_DB_Animation"
   Circle "Circle_35" at 307,299 size 12x12
      Visibility <- "10_DI_DATA_E_400_RUN"
      HorizontalMovement <- "E-400 Animation_DB_Animation"
   Circle "Circle_36" at 308,423 size 12x12
      DiagonalMovement <- "E-400 Animation_DB_Animation"
      Visibility <- "10_DI_DATA_E_400_RUN"
   Circle "Circle_37" at 357,481 size 13x13
      DiagonalMovement <- "E-400 Animation_DB_Animation"
      Visibility <- "10_DI_DATA_E_400_RUN"
   Circle "Circle_61" at 392,416 size 10x10
      DiagonalMovement <- "E-400 Animation_DB_Animation"
      Visibility <- "10_DI_DATA_E_400_RUN"
   Circle "Circle_63" at 408,416 size 10x10
      DiagonalMovement <- "E-400 Animation_DB_Animation"
      Visibility <- "10_DI_DATA_E_400_RUN"
   Circle "Circle_64" at 424,416 size 10x10
      DiagonalMovement <- "E-400 Animation_DB_Animation"
      Visibility <- "10_DI_DATA_E_400_RUN"
   Circle "Circle_65" at 456,416 size 10x10
      DiagonalMovement <- "E-400 Animation_DB_Animation"
      Visibility <- "10_DI_DATA_E_400_RUN"
   Circle "Circle_66" at 472,416 size 10x10
      DiagonalMovement <- "E-400 Animation_DB_Animation"
      Visibility <- "10_DI_DATA_E_400_RUN"
   Circle "Circle_62" at 440,416 size 10x10
      DiagonalMovement <- "E-400 Animation_DB_Animation"
      Visibility <- "10_DI_DATA_E_400_RUN"
   Circle "Circle_54" at 384,309 size 7x7
      DiagonalMovement <- "82_To_HMI_FS350 Animation"
      Visibility <- "10_DI_DATA_FS_350_FLW_OK"
   Circle "Circle_53" at 388,321 size 8x8
      DiagonalMovement <- "82_To_HMI_FS350 Animation"
      Visibility <- "10_DI_DATA_FS_350_FLW_OK"
   Circle "Circle_51" at 407,332 size 6x6
      DiagonalMovement <- "82_To_HMI_FS350 Animation"
      Visibility <- "10_DI_DATA_FS_350_FLW_OK"
   Circle "Circle_49" at 432,336 size 6x6
      DiagonalMovement <- "82_To_HMI_FS350 Animation"
      Visibility <- "10_DI_DATA_FS_350_FLW_OK"
   Circle "Circle_50" at 453,328 size 7x7
      DiagonalMovement <- "82_To_HMI_FS350 Animation"
      Visibility <- "10_DI_DATA_FS_350_FLW_OK"
   Circle "Circle_52" at 466,317 size 8x8
      DiagonalMovement <- "82_To_HMI_FS350 Animation"
      Visibility <- "10_DI_DATA_FS_350_FLW_OK"
   Circle "Circle_48" at 476,306 size 7x7
      DiagonalMovement <- "82_To_HMI_FS350 Animation"
      Visibility <- "10_DI_DATA_FS_350_FLW_OK"
   Circle "Circle_14" at 437,257 size 10x10
      DiagonalMovement <- "82_To_HMI_FS350 Animation"
      Visibility <- "10_DI_DATA_FS_350_FLW_OK"
   Circle "Circle_5" at 527,257 size 9x9
      DiagonalMovement <- "82_To_HMI_FS350 Animation"
      Visibility <- "10_DI_DATA_FS_350_FLW_OK"
   Circle "Circle_6" at 589,257 size 9x9
      DiagonalMovement <- "82_To_HMI_FS350 Animation"
      Visibility <- "10_DI_DATA_FS_350_FLW_OK"
   Circle "Circle_7" at 664,257 size 9x9
      DiagonalMovement <- "82_To_HMI_FS350 Animation"
      Visibility <- "10_DI_DATA_FS_350_FLW_OK"
   Circle "Circle_8" at 739,257 size 10x10
      DiagonalMovement <- "82_To_HMI_FS350 Animation"
      Visibility <- "10_DI_DATA_FS_350_FLW_OK"
   Circle "Circle_9" at 816,258 size 9x9
      DiagonalMovement <- "82_To_HMI_FS350 Animation"
      Visibility <- "10_DI_DATA_FS_350_FLW_OK"
   Circle "Circle_12" at 877,264 size 10x10
      Visibility <- "10_DI_DATA_FS_350_FLW_OK"
      VerticalMovement <- "82_To_HMI_FS350 Animation"
   Circle "Circle_13" at 878,359 size 10x10
      Visibility <- "10_DI_DATA_FS_350_FLW_OK"
      VerticalMovement <- "82_To_HMI_FS350 Animation"
   Circle "Circle_11" at 870,466 size 10x10
      DiagonalMovement <- "82_To_HMI_FS350 Animation"
      Visibility <- "10_DI_DATA_FS_350_FLW_OK"
   Circle "Circle_10" at 774,469 size 9x9
      DiagonalMovement <- "82_To_HMI_FS350 Animation"
      Visibility <- "10_DI_DATA_FS_350_FLW_OK"
   Circle "Circle_47" at 669,474 size 10x10
      Visibility <- "10_DI_DATA_FS_350_FLW_OK"
      VerticalMovement <- "82_To_HMI_FS350 Animation"
   Circle "Circle_46" at 667,509 size 10x10
      DiagonalMovement <- "82_To_HMI_FS350 Animation"
      Visibility <- "10_DI_DATA_FS_350_FLW_OK"
   Circle "Circle_15" at 475,635 size 10x10
      Visibility <- "10_DI_DATA_FS_350_FLW_OK"
      HorizontalMovement <- "82_To_HMI_FS350 Animation"
   Circle "Circle_16" at 518,635 size 10x10
      Visibility <- "10_DI_DATA_FS_350_FLW_OK"
      HorizontalMovement <- "82_To_HMI_FS350 Animation"
   Circle "Circle_17" at 562,635 size 10x10
      Visibility <- "10_DI_DATA_FS_350_FLW_OK"
      HorizontalMovement <- "82_To_HMI_FS350 Animation"
   Circle "Circle_18" at 661,635 size 9x9
      Visibility <- "10_DI_DATA_FS_350_FLW_OK"
      HorizontalMovement <- "82_To_HMI_FS350 Animation"
   Circle "Circle_19" at 684,635 size 9x9
      Visibility <- "10_DI_DATA_FS_350_FLW_OK"
      HorizontalMovement <- "82_To_HMI_FS350 Animation"
   Circle "Circle_21" at 403,292 size 6x6
      DiagonalMovement <- "82_To_HMI_FS350 Animation"
      Visibility <- "10_DI_DATA_FS_350_FLW_OK"
   Circle "Circle_22" at 410,301 size 6x6
      DiagonalMovement <- "82_To_HMI_FS350 Animation"
      Visibility <- "10_DI_DATA_FS_350_FLW_OK"
   Circle "Circle_25" at 418,306 size 6x6
      DiagonalMovement <- "82_To_HMI_FS350 Animation"
      Visibility <- "10_DI_DATA_FS_350_FLW_OK"
   Circle "Circle_3" at 429,307 size 7x7
      DiagonalMovement <- "82_To_HMI_FS350 Animation"
      Visibility <- "10_DI_DATA_FS_350_FLW_OK"
   Circle "Circle_4" at 445,307 size 5x5
      DiagonalMovement <- "82_To_HMI_FS350 Animation"
      Visibility <- "10_DI_DATA_FS_350_FLW_OK"
   Circle "Circle_23" at 453,302 size 5x5
      DiagonalMovement <- "82_To_HMI_FS350 Animation"
      Visibility <- "10_DI_DATA_FS_350_FLW_OK"
   Circle "Circle_24" at 460,295 size 6x6
      DiagonalMovement <- "82_To_HMI_FS350 Animation"
      Visibility <- "10_DI_DATA_FS_350_FLW_OK"
   Circle "Circle_67" at 260,764 size 8x8
      Visibility <- "10_DI_DATA_FS_332 FLW_OK"
      HorizontalMovement <- "82_To_HMI_FS332 Animation"
   Circle "Circle_68" at 411,763 size 8x8